// TIA Portal project "ESTHER_Gas_v4.0_4" (V13) (continued)
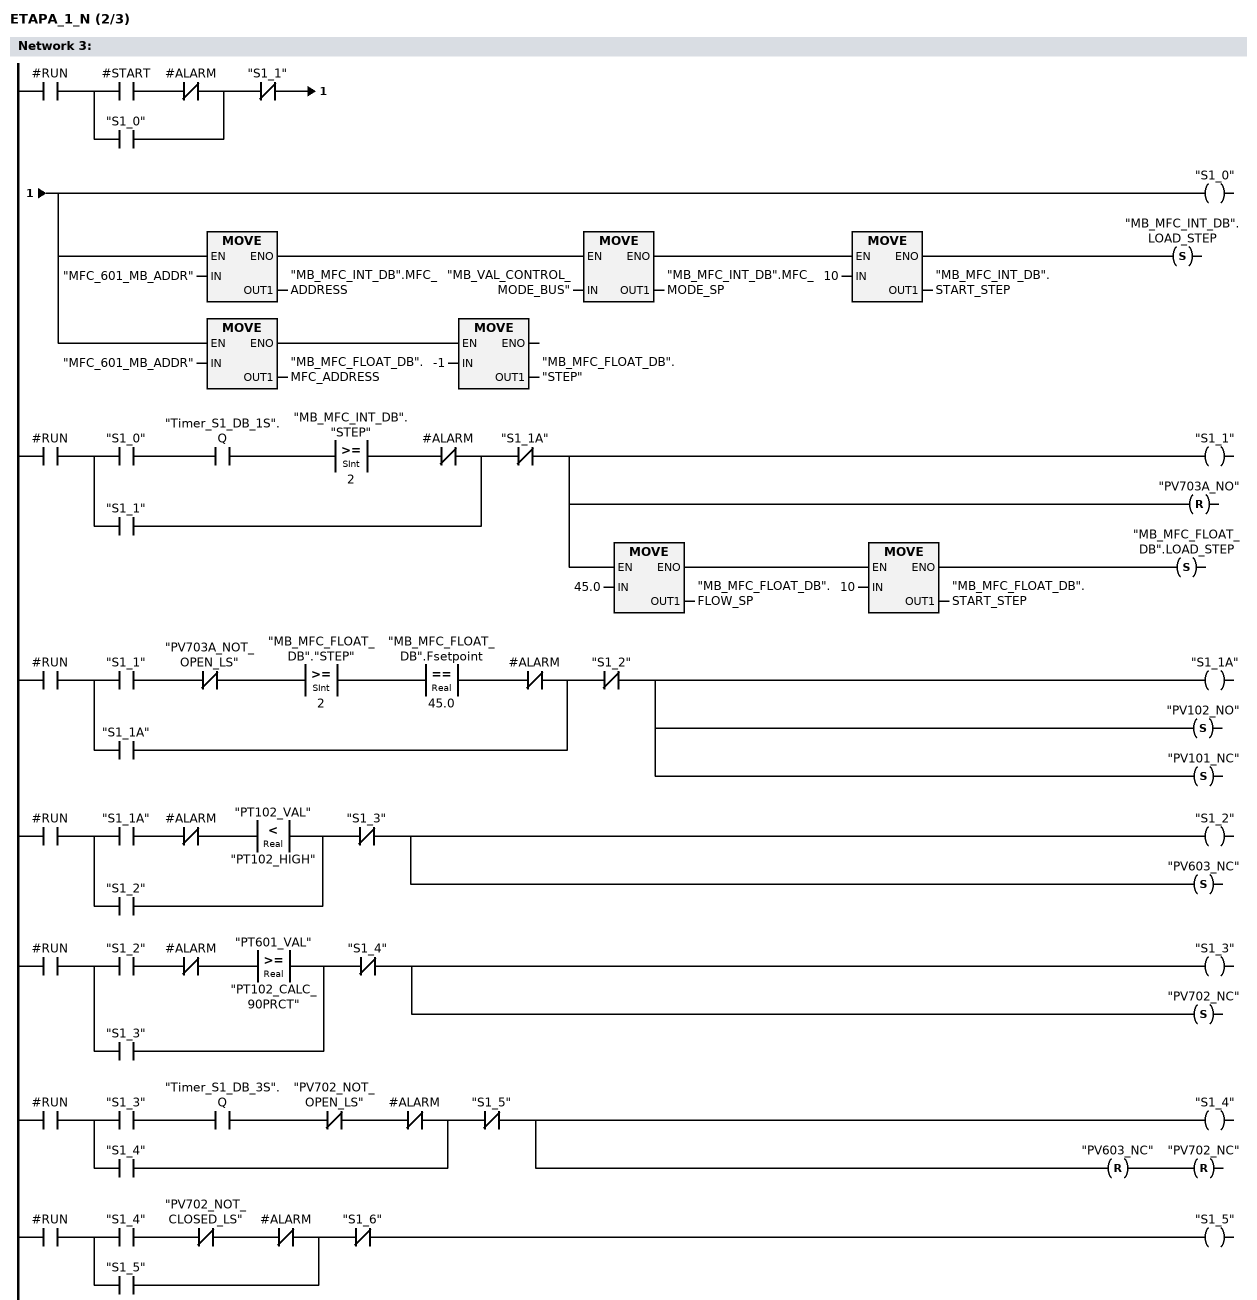
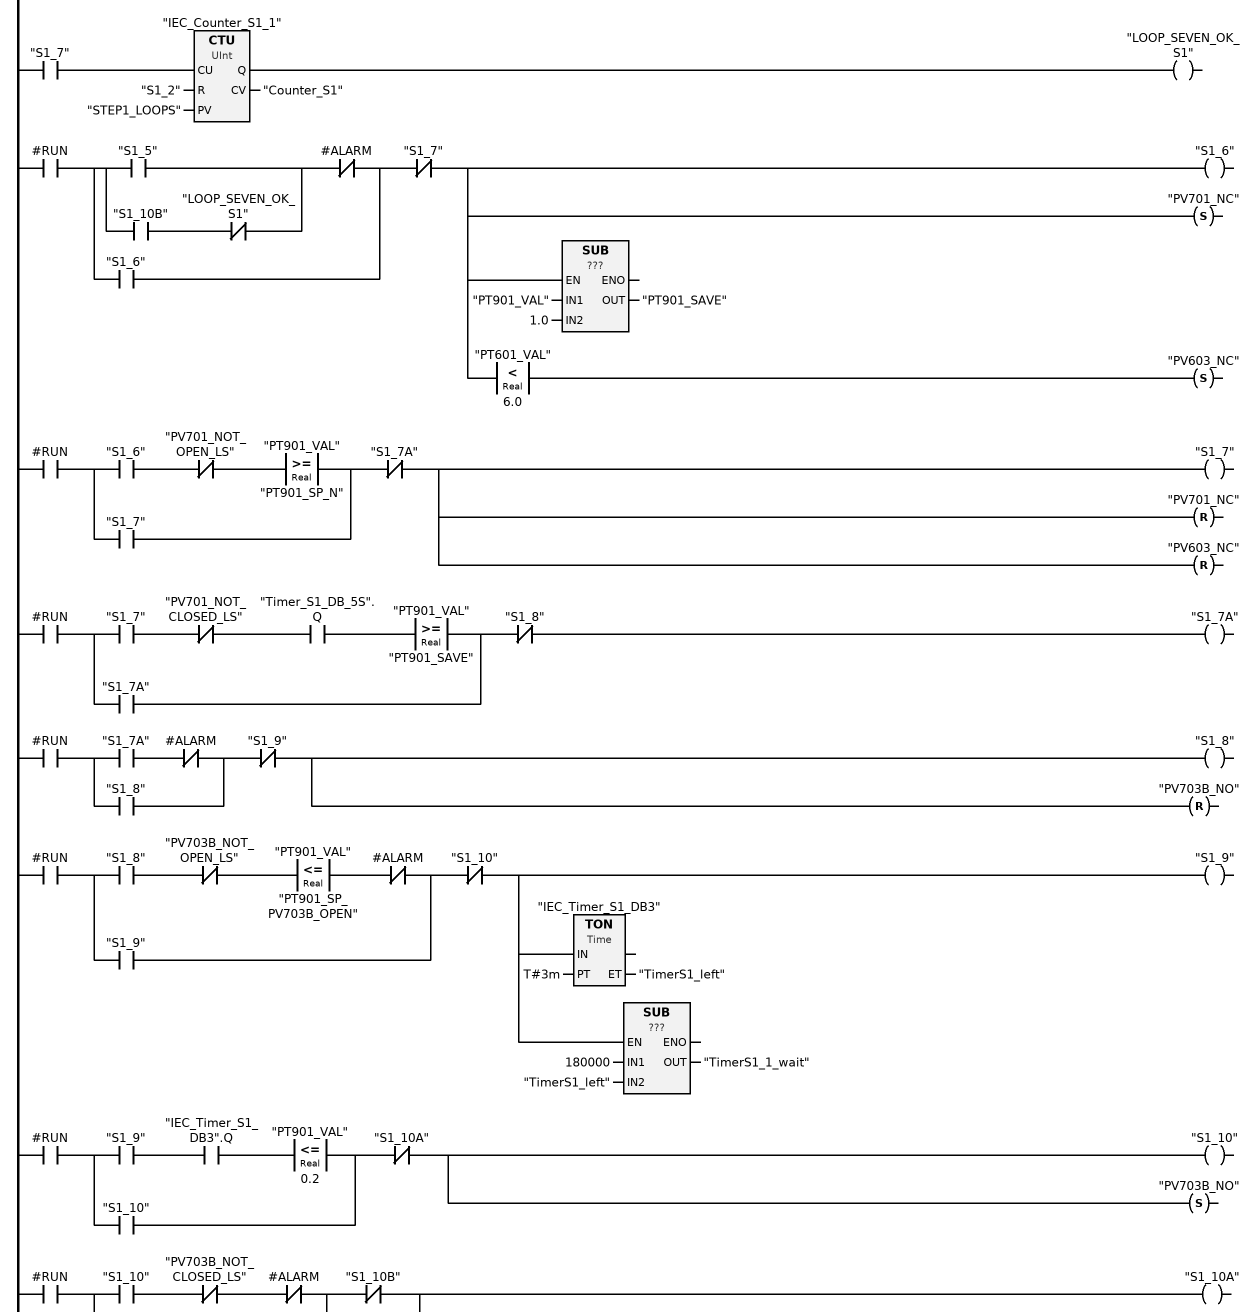
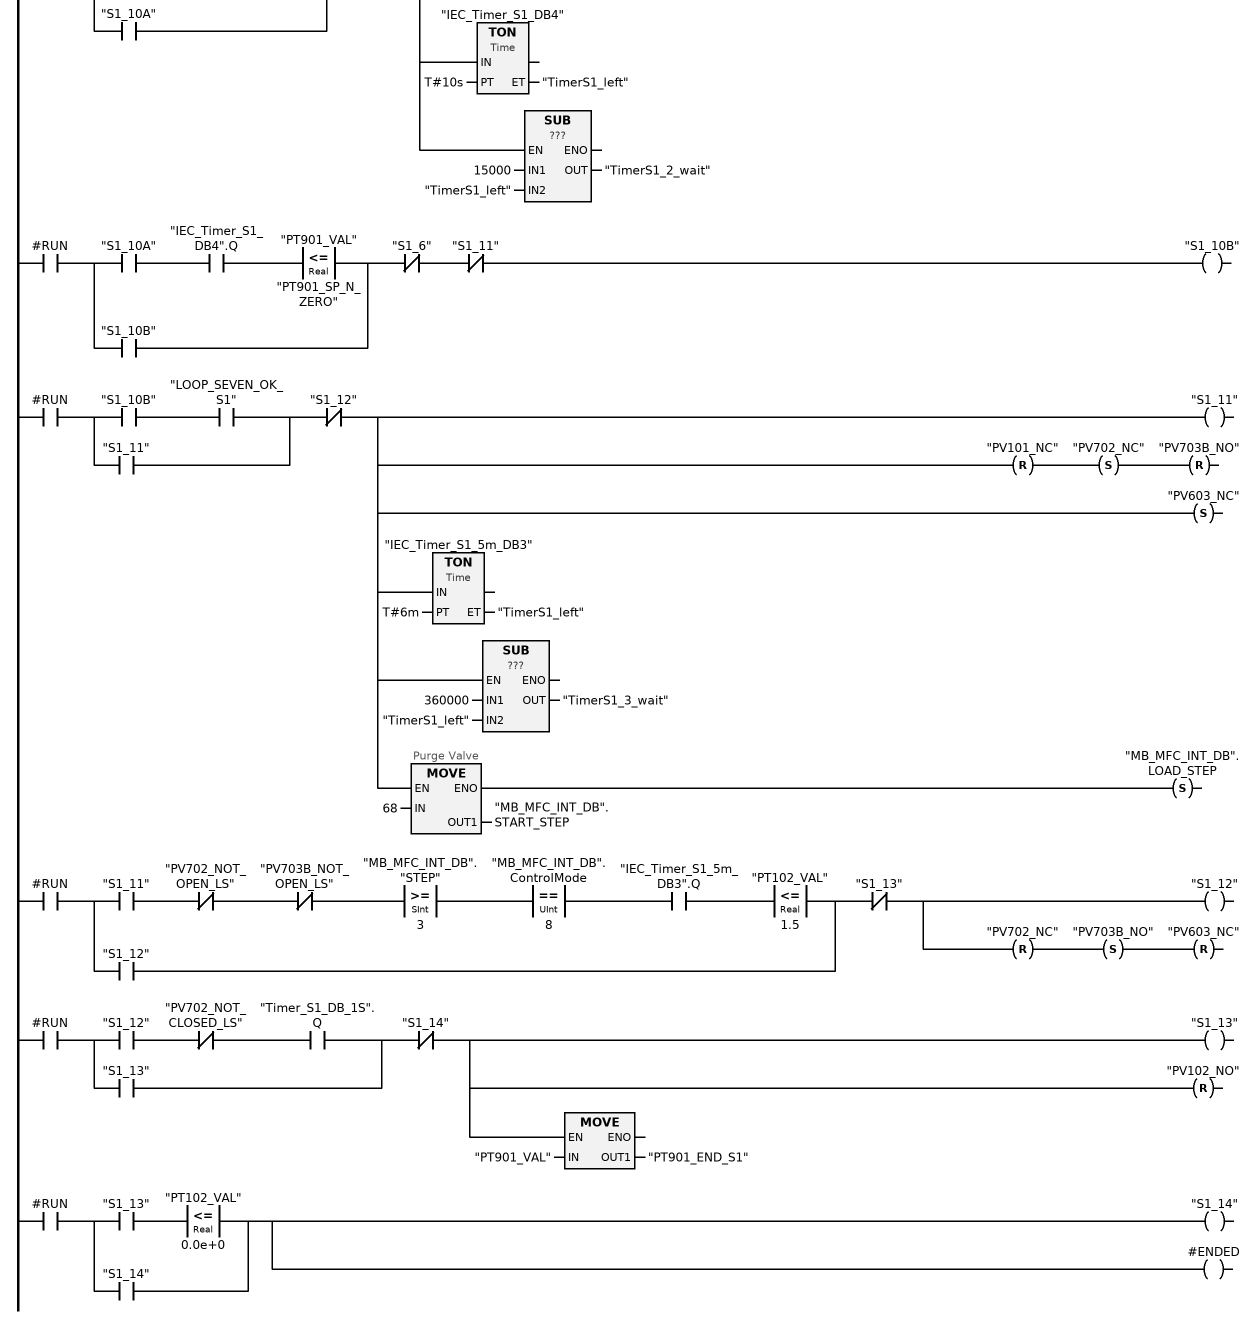
   "S1_0" := #RUN AND ((#START AND NOT #ALARM) OR "S1_0") AND NOT "S1_1";
   IF "S1_0" THEN
       "MB_MFC_INT_DB".MFC_ADDRESS := "MFC_601_MB_ADDR";
       "MB_MFC_INT_DB".MFC_MODE_SP := "MB_VAL_CONTROL_MODE_BUS";
       "MB_MFC_INT_DB".START_STEP := 10;
       "MB_MFC_INT_DB".LOAD_STEP := TRUE;
       "MB_MFC_FLOAT_DB".MFC_ADDRESS := "MFC_601_MB_ADDR";
       "MB_MFC_FLOAT_DB"."STEP" := -1;
   END_IF;
   "S1_1" := #RUN AND (("S1_0" AND "Timer_S1_DB_1S".Q AND ("MB_MFC_INT_DB"."STEP" >= 2) AND NOT #ALARM) OR "S1_1") AND NOT "S1_1A";
   IF "S1_1" THEN
       "PV703A_NO" := FALSE;
       "MB_MFC_FLOAT_DB".FLOW_SP := 45.0;
       "MB_MFC_FLOAT_DB".START_STEP := 10;
       "MB_MFC_FLOAT_DB".LOAD_STEP := TRUE;
   END_IF;
   "S1_1A" := #RUN AND (("S1_1" AND NOT "PV703A_NOT_OPEN_LS" AND ("MB_MFC_FLOAT_DB"."STEP" >= 2) AND ("MB_MFC_FLOAT_DB".Fsetpoint = 45.0) AND NOT #ALARM) OR "S1_1A") AND NOT "S1_2";
   IF "S1_1A" THEN
       "PV102_NO" := TRUE;
       "PV101_NC" := TRUE;
   END_IF;
   "S1_2" := #RUN AND (("S1_1A" AND NOT #ALARM AND ("PT102_VAL" < "PT102_HIGH")) OR "S1_2") AND NOT "S1_3";
   IF "S1_2" THEN "PV603_NC" := TRUE; END_IF;
   "S1_3" := #RUN AND (("S1_2" AND NOT #ALARM AND ("PT601_VAL" >= "PT102_CALC_90PRCT")) OR "S1_3") AND NOT "S1_4";
   IF "S1_3" THEN "PV702_NC" := TRUE; END_IF;
   "S1_4" := #RUN AND (("S1_3" AND "Timer_S1_DB_3S".Q AND NOT "PV702_NOT_OPEN_LS" AND NOT #ALARM) OR "S1_4") AND NOT "S1_5";
   IF "S1_4" THEN
       "PV603_NC" := FALSE;
       "PV702_NC" := FALSE;
   END_IF;
   "S1_5" := #RUN AND (("S1_4" AND NOT "PV702_NOT_CLOSED_LS" AND NOT #ALARM) OR "S1_5") AND NOT "S1_6";
   "IEC_Counter_S1_1".CTU(CU := "S1_7", R := "S1_2", PV := "STEP1_LOOPS", CV => "Counter_S1");
   "LOOP_SEVEN_OK_S1" := "IEC_Counter_S1_1".Q;
   "S1_6" := #RUN AND ((("S1_5" OR ("S1_10B" AND NOT "LOOP_SEVEN_OK_S1")) AND NOT #ALARM) OR "S1_6") AND NOT "S1_7";
   IF "S1_6" THEN
       "PV701_NC" := TRUE;
       "PT901_SAVE" := "PT901_VAL" - 1.0;
   END_IF;
   IF "S1_6" AND ("PT601_VAL" < 6.0) THEN "PV603_NC" := TRUE; END_IF;
   "S1_7" := #RUN AND (("S1_6" AND NOT "PV701_NOT_OPEN_LS" AND ("PT901_VAL" >= "PT901_SP_N")) OR "S1_7") AND NOT "S1_7A";
   IF "S1_7" THEN
       "PV701_NC" := FALSE;
       "PV603_NC" := FALSE;
   END_IF;
   "S1_7A" := #RUN AND (("S1_7" AND NOT "PV701_NOT_CLOSED_LS" AND "Timer_S1_DB_5S".Q AND ("PT901_VAL" >= "PT901_SAVE")) OR "S1_7A") AND NOT "S1_8";
   "S1_8" := #RUN AND (("S1_7A" AND NOT #ALARM) OR "S1_8") AND NOT "S1_9";
   IF "S1_8" THEN "PV703B_NO" := FALSE; END_IF;
   "S1_9" := #RUN AND (("S1_8" AND NOT "PV703B_NOT_OPEN_LS" AND ("PT901_VAL" <= "PT901_SP_PV703B_OPEN") AND NOT #ALARM) OR "S1_9") AND NOT "S1_10";
   "IEC_Timer_S1_DB3".TON(IN := "S1_9", PT := T#3m, ET => "TimerS1_left");
   IF "S1_9" THEN "TimerS1_1_wait" := 180000 - "TimerS1_left"; END_IF;
   "S1_10" := #RUN AND (("S1_9" AND "IEC_Timer_S1_DB3".Q AND ("PT901_VAL" <= 0.2)) OR "S1_10") AND NOT "S1_10A";
   IF "S1_10" THEN "PV703B_NO" := TRUE; END_IF;
   "S1_10A" := #RUN AND (("S1_10" AND NOT "PV703B_NOT_CLOSED_LS" AND NOT #ALARM) OR "S1_10A") AND NOT "S1_10B";
   "IEC_Timer_S1_DB4".TON(IN := "S1_10A", PT := T#10s, ET => "TimerS1_left");
   IF "S1_10A" THEN "TimerS1_2_wait" := 15000 - "TimerS1_left"; END_IF;
   "S1_10B" := #RUN AND (("S1_10A" AND "IEC_Timer_S1_DB4".Q AND ("PT901_VAL" <= "PT901_SP_N_ZERO")) OR "S1_10B") AND NOT "S1_6" AND NOT "S1_11";
   "S1_11" := #RUN AND (("S1_10B" AND "LOOP_SEVEN_OK_S1") OR "S1_11") AND NOT "S1_12";
   IF "S1_11" THEN
       "PV101_NC" := FALSE;
       "PV702_NC" := TRUE;
       "PV703B_NO" := FALSE;
       "PV603_NC" := TRUE;
   END_IF;
   "IEC_Timer_S1_5m_DB3".TON(IN := "S1_11", PT := T#6m, ET => "TimerS1_left");
   IF "S1_11" THEN
       "TimerS1_3_wait" := 360000 - "TimerS1_left";
       "MB_MFC_INT_DB".START_STEP := 68;   // Purge Valve
       "MB_MFC_INT_DB".LOAD_STEP := TRUE;
   END_IF;
   "S1_12" := #RUN AND (("S1_11" AND NOT "PV702_NOT_OPEN_LS" AND NOT "PV703B_NOT_OPEN_LS" AND ("MB_MFC_INT_DB"."STEP" >= 3) AND ("MB_MFC_INT_DB".ControlMode = 8) AND "IEC_Timer_S1_5m_DB3".Q AND ("PT102_VAL" <= 1.5)) OR "S1_12") AND NOT "S1_13";
   IF "S1_12" THEN
       "PV702_NC" := FALSE;
       "PV703B_NO" := TRUE;
       "PV603_NC" := FALSE;
   END_IF;
   "S1_13" := #RUN AND (("S1_12" AND NOT "PV702_NOT_CLOSED_LS" AND "Timer_S1_DB_1S".Q) OR "S1_13") AND NOT "S1_14";
   IF "S1_13" THEN
       "PV102_NO" := FALSE;
       "PT901_END_S1" := "PT901_VAL";
   END_IF;
   "S1_14" := #RUN AND (("S1_13" AND ("PT102_VAL" <= 0.0e+0)) OR "S1_14");
   #ENDED := "S1_14";
END_REGION

REGION Network 4
   // Timers
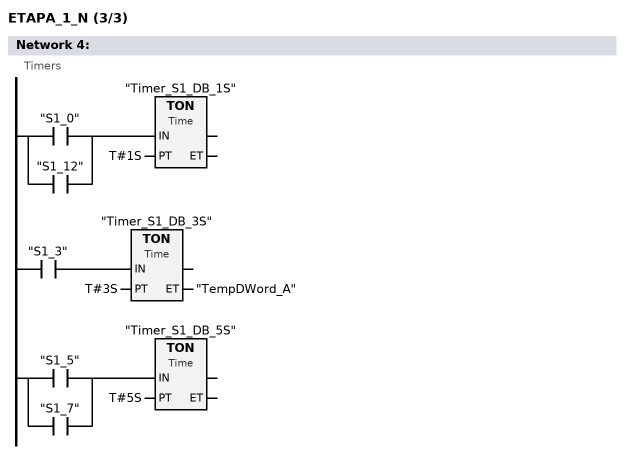
   "Timer_S1_DB_1S".TON(IN := "S1_0" OR "S1_12", PT := T#1S);
   "Timer_S1_DB_3S".TON(IN := "S1_3", PT := T#3S, ET => "TempDWord_A");
   "Timer_S1_DB_5S".TON(IN := "S1_5" OR "S1_7", PT := T#5S);
END_REGION

REGION Network 5: NC Temp
END_REGION
END_FUNCTION

FUNCTION "ETAPA_2" : Void   // FC2, LAD
{ S7_Optimized_Access := 'FALSE' }
VERSION : 0.1
// Varrimento com HELIO 1
   VAR_TEMP   // added for the SCL form of the ladder/FBD networks
      _w1 : Bool;
   END_VAR
BEGIN

REGION Network 1
   // Alarm Set points of this step
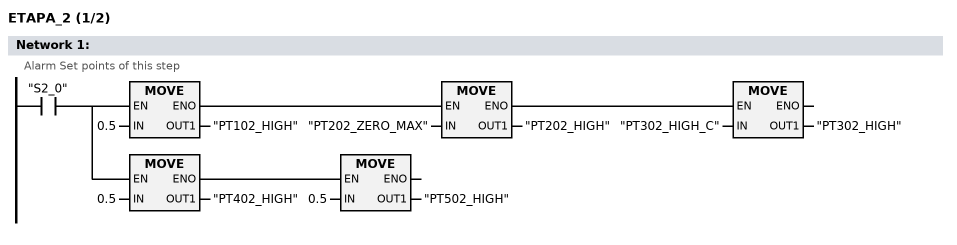
   RUNG wire#powerrail
      Contact( "S2_0" )
      wire#w1
      { S7_GenerateENO := "TRUE" } Move(in := 0.5, out1 => "PT102_HIGH")
      { S7_GenerateENO := "TRUE" } Move(in := "PT202_ZERO_MAX", out1 => "PT202_HIGH")
      { S7_GenerateENO := "TRUE" } Move(in := "PT302_HIGH_C", out1 => "PT302_HIGH")
   END_RUNG
   RUNG wire#w1
      { S7_GenerateENO := "TRUE" } Move(in := 0.5, out1 => "PT402_HIGH")
      { S7_GenerateENO := "TRUE" } Move(in := 0.5, out1 => "PT502_HIGH")
   END_RUNG
   // the same network as SCL:
   // ENO of a box is taken as its EN; it also drops when the box reports an error
   IF "S2_0" THEN
       "PT102_HIGH" := 0.5;
       "PT202_HIGH" := "PT202_ZERO_MAX";
       "PT302_HIGH" := "PT302_HIGH_C";
       "PT402_HIGH" := 0.5;
       "PT502_HIGH" := 0.5;
   END_IF;
END_REGION

REGION Network 2
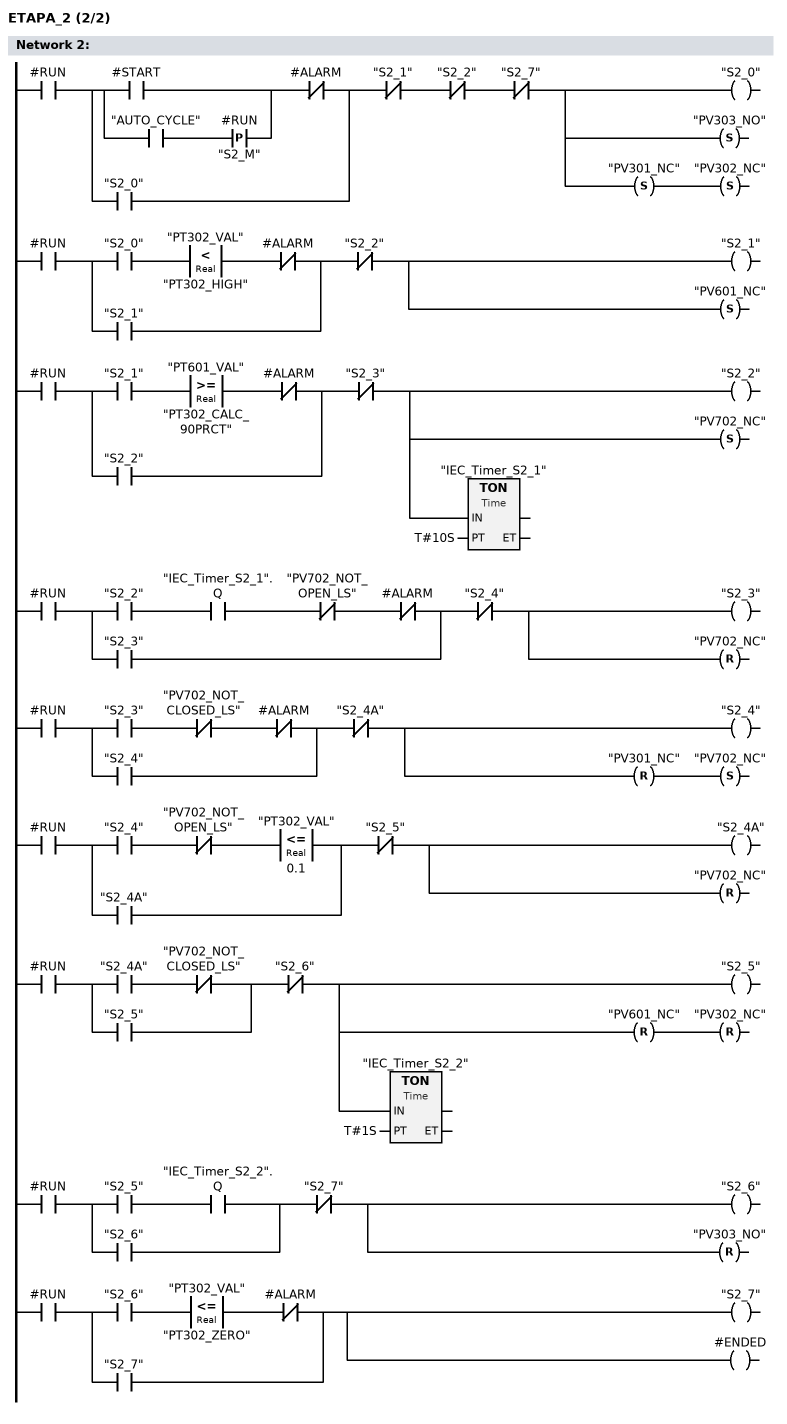
   #_w1 := #RUN AND "AUTO_CYCLE" AND #RUN AND NOT "S2_M";   // rising edge of #RUN
   "S2_M" := #RUN;
   "S2_0" := ((((#RUN AND #START) OR #_w1) AND NOT #ALARM) OR (#RUN AND "S2_0")) AND NOT "S2_1" AND NOT "S2_2" AND NOT "S2_7";
   IF "S2_0" THEN
       "PV303_NO" := TRUE;
       "PV301_NC" := TRUE;
       "PV302_NC" := TRUE;
   END_IF;
   "S2_1" := #RUN AND (("S2_0" AND ("PT302_VAL" < "PT302_HIGH") AND NOT #ALARM) OR "S2_1") AND NOT "S2_2";
   IF "S2_1" THEN "PV601_NC" := TRUE; END_IF;
   "S2_2" := #RUN AND (("S2_1" AND ("PT601_VAL" >= "PT302_CALC_90PRCT") AND NOT #ALARM) OR "S2_2") AND NOT "S2_3";
   IF "S2_2" THEN "PV702_NC" := TRUE; END_IF;
   "IEC_Timer_S2_1".TON(IN := "S2_2", PT := T#10S);
   "S2_3" := #RUN AND (("S2_2" AND "IEC_Timer_S2_1".Q AND NOT "PV702_NOT_OPEN_LS" AND NOT #ALARM) OR "S2_3") AND NOT "S2_4";
   IF "S2_3" THEN "PV702_NC" := FALSE; END_IF;
   "S2_4" := #RUN AND (("S2_3" AND NOT "PV702_NOT_CLOSED_LS" AND NOT #ALARM) OR "S2_4") AND NOT "S2_4A";
   IF "S2_4" THEN
       "PV301_NC" := FALSE;
       "PV702_NC" := TRUE;
   END_IF;
   "S2_4A" := #RUN AND (("S2_4" AND NOT "PV702_NOT_OPEN_LS" AND ("PT302_VAL" <= 0.1)) OR "S2_4A") AND NOT "S2_5";
   IF "S2_4A" THEN "PV702_NC" := FALSE; END_IF;
   "S2_5" := #RUN AND (("S2_4A" AND NOT "PV702_NOT_CLOSED_LS") OR "S2_5") AND NOT "S2_6";
   IF "S2_5" THEN
       "PV601_NC" := FALSE;
       "PV302_NC" := FALSE;
   END_IF;
   "IEC_Timer_S2_2".TON(IN := "S2_5", PT := T#1S);
   "S2_6" := #RUN AND (("S2_5" AND "IEC_Timer_S2_2".Q) OR "S2_6") AND NOT "S2_7";
   IF "S2_6" THEN "PV303_NO" := FALSE; END_IF;
   "S2_7" := #RUN AND (("S2_6" AND ("PT302_VAL" <= "PT302_ZERO") AND NOT #ALARM) OR "S2_7");
   #ENDED := "S2_7";
END_REGION
END_FUNCTION

FUNCTION "ETAPA_0" : Void   // FC3, LAD
{ S7_Optimized_Access := 'FALSE' }
VERSION : 0.1
// ETAPA 0 - ESTADO STAND-BY
   VAR_TEMP   // added for the SCL form of the ladder/FBD networks
      _w1 : Bool;
      _w2 : Bool;
   END_VAR
BEGIN

REGION Network 1
   // PT Alarm  Set Points
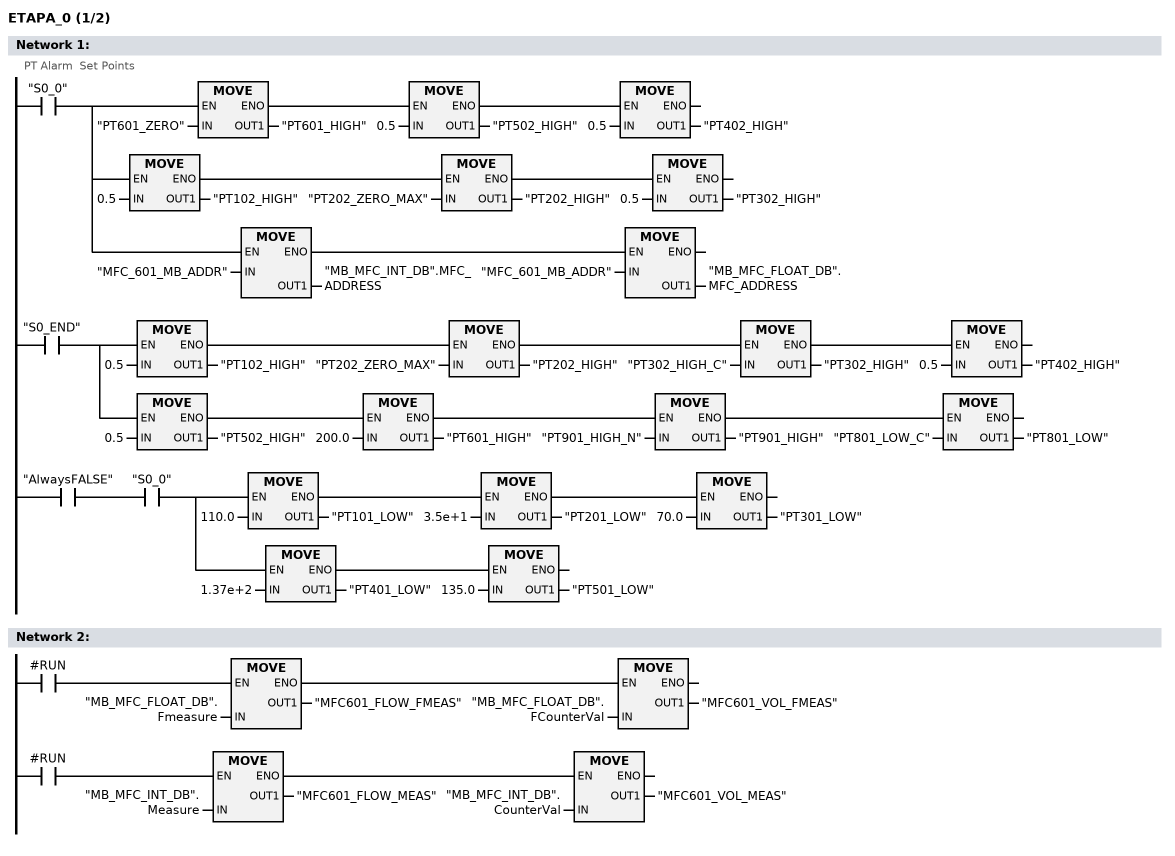
   RUNG wire#powerrail
      Contact( "S0_0" )
      wire#w1
      { S7_GenerateENO := "TRUE" } Move(in := "PT601_ZERO", out1 => "PT601_HIGH")
      { S7_GenerateENO := "TRUE" } Move(in := 0.5, out1 => "PT502_HIGH")
      { S7_GenerateENO := "TRUE" } Move(in := 0.5, out1 => "PT402_HIGH")
   END_RUNG
   RUNG wire#w1
      { S7_GenerateENO := "TRUE" } Move(in := 0.5, out1 => "PT102_HIGH")
      { S7_GenerateENO := "TRUE" } Move(in := "PT202_ZERO_MAX", out1 => "PT202_HIGH")
      { S7_GenerateENO := "TRUE" } Move(in := 0.5, out1 => "PT302_HIGH")
   END_RUNG
   RUNG wire#w1
      Move(in := "MFC_601_MB_ADDR", out1 => "MB_MFC_INT_DB".MFC_ADDRESS)
      Move(in := "MFC_601_MB_ADDR", out1 => "MB_MFC_FLOAT_DB".MFC_ADDRESS)
   END_RUNG
   RUNG wire#powerrail
      Contact( "S0_END" )
      wire#w2
      { S7_GenerateENO := "TRUE" } Move(in := 0.5, out1 => "PT102_HIGH")
      { S7_GenerateENO := "TRUE" } Move(in := "PT202_ZERO_MAX", out1 => "PT202_HIGH")
      { S7_GenerateENO := "TRUE" } Move(in := "PT302_HIGH_C", out1 => "PT302_HIGH")
      { S7_GenerateENO := "TRUE" } Move(in := 0.5, out1 => "PT402_HIGH")
   END_RUNG
   RUNG wire#w2
      { S7_GenerateENO := "TRUE" } Move(in := 0.5, out1 => "PT502_HIGH")
      { S7_GenerateENO := "TRUE" } Move(in := 200.0, out1 => "PT601_HIGH")
      { S7_GenerateENO := "TRUE" } Move(in := "PT901_HIGH_N", out1 => "PT901_HIGH")
      { S7_GenerateENO := "TRUE" } Move(in := "PT801_LOW_C", out1 => "PT801_LOW")
   END_RUNG
   RUNG wire#powerrail
      Contact( "AlwaysFALSE" )
      Contact( "S0_0" )
      wire#w3
      { S7_GenerateENO := "TRUE" } Move(in := 110.0, out1 => "PT101_LOW")
      { S7_GenerateENO := "TRUE" } Move(in := 3.5e+1, out1 => "PT201_LOW")
      { S7_GenerateENO := "TRUE" } Move(in := 70.0, out1 => "PT301_LOW")
   END_RUNG
   RUNG wire#w3
      { S7_GenerateENO := "TRUE" } Move(in := 1.37e+2, out1 => "PT401_LOW")
      { S7_GenerateENO := "TRUE" } Move(in := 135.0, out1 => "PT501_LOW")
   END_RUNG
   // the same network as SCL:
   // ENO of a box is taken as its EN; it also drops when the box reports an error
   IF "S0_0" THEN
       "PT601_HIGH" := "PT601_ZERO";
       "PT502_HIGH" := 0.5;
       "PT402_HIGH" := 0.5;
       "PT102_HIGH" := 0.5;
       "PT202_HIGH" := "PT202_ZERO_MAX";
       "PT302_HIGH" := 0.5;
       "MB_MFC_INT_DB".MFC_ADDRESS := "MFC_601_MB_ADDR";
       "MB_MFC_FLOAT_DB".MFC_ADDRESS := "MFC_601_MB_ADDR";
   END_IF;
   IF "S0_END" THEN
       "PT102_HIGH" := 0.5;
       "PT202_HIGH" := "PT202_ZERO_MAX";
       "PT302_HIGH" := "PT302_HIGH_C";
       "PT402_HIGH" := 0.5;
       "PT502_HIGH" := 0.5;
       "PT601_HIGH" := 200.0;
       "PT901_HIGH" := "PT901_HIGH_N";
       "PT801_LOW" := "PT801_LOW_C";
   END_IF;
   IF "AlwaysFALSE" AND "S0_0" THEN
       "PT101_LOW" := 110.0;
       "PT201_LOW" := 3.5e+1;
       "PT301_LOW" := 70.0;
       "PT401_LOW" := 1.37e+2;
       "PT501_LOW" := 135.0;
   END_IF;
END_REGION

REGION Network 2
   RUNG wire#powerrail
      Contact( #RUN )
      { S7_GenerateENO := "TRUE" } Move(in := "MB_MFC_FLOAT_DB".Fmeasure, out1 => "MFC601_FLOW_FMEAS")
      { S7_GenerateENO := "TRUE" } Move(in := "MB_MFC_FLOAT_DB".FCounterVal, out1 => "MFC601_VOL_FMEAS")
   END_RUNG
   RUNG wire#powerrail
      Contact( #RUN )
      { S7_GenerateENO := "TRUE" } Move(in := "MB_MFC_INT_DB".Measure, out1 => "MFC601_FLOW_MEAS")
      { S7_GenerateENO := "TRUE" } Move(in := "MB_MFC_INT_DB".CounterVal, out1 => "MFC601_VOL_MEAS")
   END_RUNG
   // the same network as SCL:
   // ENO of a box is taken as its EN; it also drops when the box reports an error
   IF #RUN THEN
       "MFC601_FLOW_FMEAS" := "MB_MFC_FLOAT_DB".Fmeasure;
       "MFC601_VOL_FMEAS" := "MB_MFC_FLOAT_DB".FCounterVal;
       "MFC601_FLOW_MEAS" := "MB_MFC_INT_DB".Measure;
       "MFC601_VOL_MEAS" := "MB_MFC_INT_DB".CounterVal;
   END_IF;
END_REGION

REGION Network 3
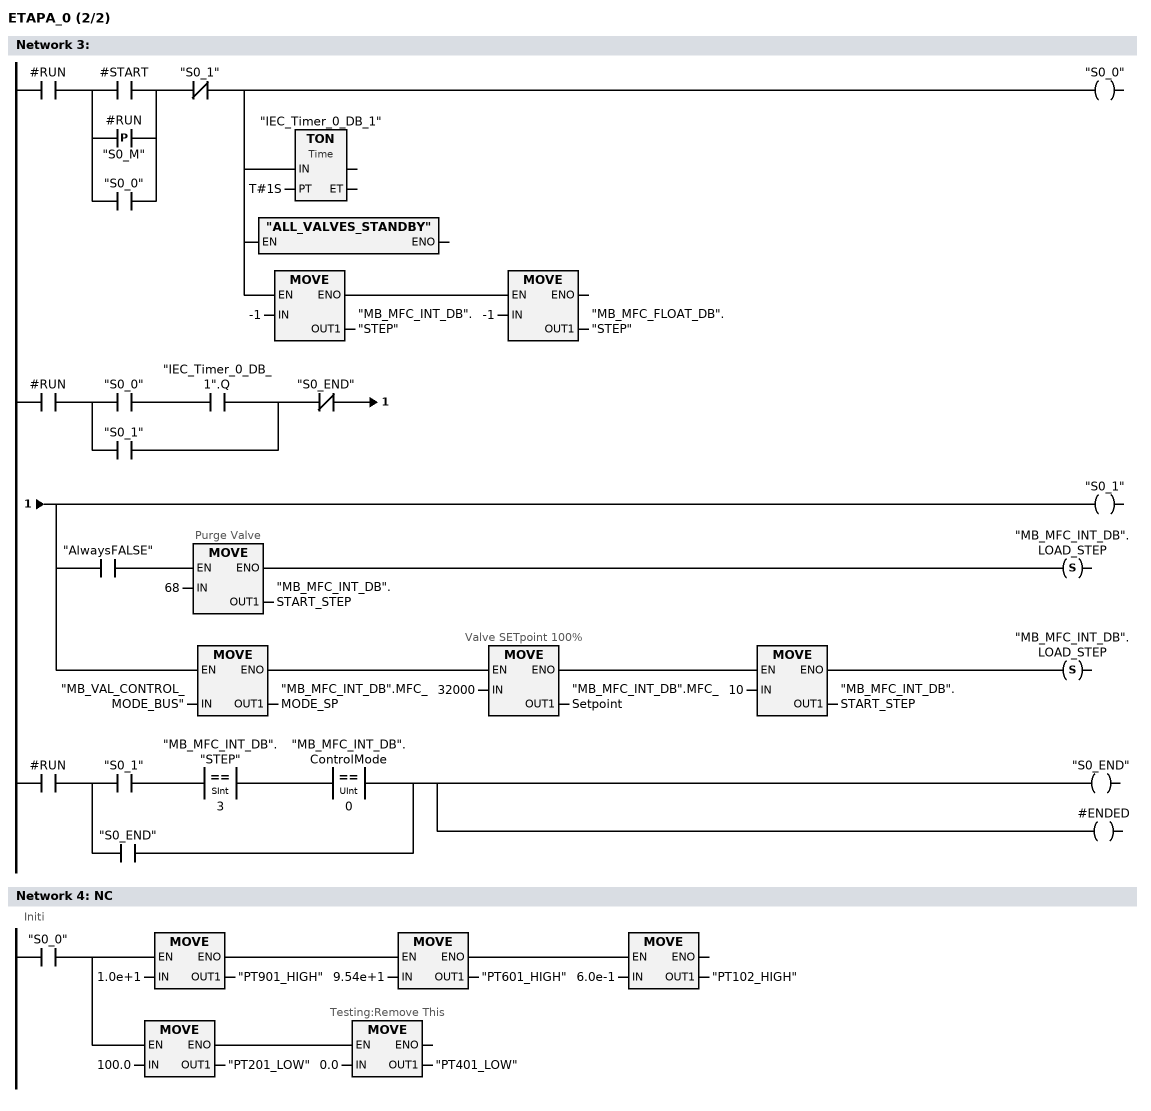
   #_w1 := #RUN AND #RUN AND NOT "S0_M";   // rising edge of #RUN
   "S0_M" := #RUN;
   "S0_0" := ((#RUN AND #START) OR #_w1 OR (#RUN AND "S0_0")) AND NOT "S0_1";
   "IEC_Timer_0_DB_1".TON(IN := "S0_0", PT := T#1S);
   #_w2 := "S0_0";
   IF #_w2 THEN
       "ALL_VALVES_STANDBY"();
       "MB_MFC_INT_DB"."STEP" := -1;
       "MB_MFC_FLOAT_DB"."STEP" := -1;
   END_IF;
   "S0_1" := #RUN AND (("S0_0" AND "IEC_Timer_0_DB_1".Q) OR "S0_1") AND NOT "S0_END";
   IF "S0_1" AND "AlwaysFALSE" THEN
       "MB_MFC_INT_DB".START_STEP := 68;   // Purge Valve
       "MB_MFC_INT_DB".LOAD_STEP := TRUE;
   END_IF;
   IF "S0_1" THEN
       "MB_MFC_INT_DB".MFC_MODE_SP := "MB_VAL_CONTROL_MODE_BUS";
       "MB_MFC_INT_DB".MFC_Setpoint := 32000;   // Valve SETpoint 100%
       "MB_MFC_INT_DB".START_STEP := 10;
       "MB_MFC_INT_DB".LOAD_STEP := TRUE;
   END_IF;
   "S0_END" := #RUN AND (("S0_1" AND ("MB_MFC_INT_DB"."STEP" = 3) AND ("MB_MFC_INT_DB".ControlMode = 0)) OR "S0_END");
   #ENDED := "S0_END";
END_REGION

REGION Network 4: NC
   // Initi
   RUNG wire#powerrail
      Contact( "S0_0" )
      wire#w1
      { S7_GenerateENO := "TRUE" } Move(in := 1.0e+1, out1 => "PT901_HIGH")
      { S7_GenerateENO := "TRUE" } Move(in := 9.54e+1, out1 => "PT601_HIGH")
      { S7_GenerateENO := "TRUE" } Move(in := 6.0e-1, out1 => "PT102_HIGH")
   END_RUNG
   RUNG wire#w1
      { S7_GenerateENO := "TRUE" } Move(in := 100.0, out1 => "PT201_LOW")
      { S7_GenerateENO := "TRUE" } Move(in := 0.0, out1 => "PT401_LOW")   // Testing:Remove This
   END_RUNG
   // the same network as SCL:
   // ENO of a box is taken as its EN; it also drops when the box reports an error
   IF "S0_0" THEN
       "PT901_HIGH" := 1.0e+1;
       "PT601_HIGH" := 9.54e+1;
       "PT102_HIGH" := 6.0e-1;
       "PT201_LOW" := 100.0;
       "PT401_LOW" := 0.0;   // Testing:Remove This
   END_IF;
END_REGION
END_FUNCTION

FUNCTION "ETAPA_3" : Void   // FC4, LAD
{ S7_Optimized_Access := 'FALSE' }
VERSION : 0.1
// Injeção de Oxigénio
   VAR_TEMP   // added for the SCL form of the ladder/FBD networks
      _w1 : Bool;
   END_VAR
BEGIN

REGION Network 1
   // Alarm Set Points
